DATA_BLOCK "DB_COM_REC_AUX"   // DB37
{ S7_Optimized_Access := 'FALSE' }
VERSION : 0.1
   VAR
      x : Bool;   // Ninguna bomba de intercambiador de soplado en marcha
      x1 : Bool;   // Ninguna bomba de chillers de soplado en marcha
      x2 : Bool;   // Ninguna bomba de intercambiador de envasado en marcha
      x3 : Bool;   // Ninguna bomba de chillers de envasado en marcha
      x4 : Bool;   // Ninguna bomba de torre de enfiamiento de chillers en marcha
      x5 : Bool;   // Ningún Chiller de soplado habilitado
      x6 : Bool;   // Ningún chiller de envasado habilitado
      x7 : Bool;   // Alarma Presente en Chiller de soplado Grande
      x8 : Bool;   // Alarma Presente en Chiller de envasado Grande
      x9 : Bool;   // Chiller de soplado Grande en su máxima capacidad
      x10 : Bool;   // Chiller de envasado Grande en su máxima capacidad
      x11 : Bool;   // Falla Térmico MT007
      x12 : Bool;   // Falla Contactor MT007
      x13 : Bool;   // Falla Térmico MT008
      x14 : Bool;   // Falla Contactor MT008
      x15 : Bool;   // Falla Térmico MT009
      x16 : Bool;   // Falla Contactor MT009
      x17 : Bool;   // Falla Térmico MT010
      x18 : Bool;   // Falla Contactor MT010
      x19 : Bool;   // Falla Térmico MP010
      x20 : Bool;   // Falla Contactor MP010
      x21 : Bool;   // Falla Térmico MP011
      x22 : Bool;   // Falla Contactor MP011
      x23 : Bool;   // Falla Térmico MP012
      x24 : Bool;   // Falla Contactor MP012
      x25 : Bool;   // Falla Térmico MP013
      x26 : Bool;   // Falla Contactor MP013
      x27 : Bool;   // Falla Térmico MP018
      x28 : Bool;   // Falla Contactor MP018
      x29 : Bool;   // Falla Térmico MP019
      x30 : Bool;   // Falla Contactor MP019
      x31 : Bool;   // Falla Térmico V001
      x32 : Bool;   // Falla Contactor V001
      x33 : Bool;   // Falla Térmico V002
      x34 : Bool;   // Falla Contactor V002
      x35 : Bool;   // Falla Térmico V003
      x36 : Bool;   // Falla Contactor V003
      x37 : Bool;   // Falla Térmico MC060
      x38 : Bool;   // Falla Contactor MC060
      x39 : Bool;   // Falla Térmico MC061
      x40 : Bool;   // Falla Contactor MC061
      x41 : Bool;   // Falla Térmico MC062
      x42 : Bool;   // Falla Contactor MC062
      x43 : Bool;   // Falla Térmico MC063
      x44 : Bool;   // Falla Contactor MC063
      x45 : Bool;   // Falla Térmico MC064
      x46 : Bool;   // Falla Contactor MC064
      x47 : Bool;   // Falla Térmico MS050
      x48 : Bool;   // Falla Contactor MS050
      x49 : Bool;   // Falla Térmico MS051
      x50 : Bool;   // Falla Contactor MS051
      x51 : Bool;   // Falla Térmico MS052
      x52 : Bool;   // Falla Contactor MS052
      x53 : Bool;   // Falla Térmico MS053
      x54 : Bool;   // Falla Contactor MS053
      x55 : Bool;   // Falla Presostato Chillers
      x56 : Bool;   // Falla Térmico MS054
      x57 : Bool;   // Falla Contactor MS054
      x58 : Bool;   // Falla Térmico MS055
      x59 : Bool;   // Falla Contactor MS055
      x60 : Bool;   // Falla Térmico MV030
      x61 : Bool;   // Falla Contactor MV030
      x62 : Bool;   // Falla Térmico MV031
      x63 : Bool;   // Falla Contactor MV031
      x64 : Bool;   // Falla Térmico MP014
      x65 : Bool;   // Falla Contactor MP014
      x66 : Bool;   // Falla Térmico MP015
      x67 : Bool;   // Falla Contactor MP015
      x68 : Bool;   // Falla Térmico MC001
      x69 : Bool;   // Falla Contactor MC001
      x70 : Bool;   // Falla Térmico MC002
      x71 : Bool;   // Falla Contactor MC002
      x72 : Bool;   // Falla Térmico MC003
      x73 : Bool;   // Falla Contactor MC003
      x74 : Bool;   // Falla Térmico MC004
      x75 : Bool;   // Falla Contactor MC004
      x76 : Bool;   // Falla Térmico MC005
      x77 : Bool;   // Falla Contactor MC005
      x78 : Bool;   // Falla Flujostato Torres Cavaleto
      x79 : Bool;   // Falla Compresor ABC2 Baja Presion de Aceite
      x80 : Bool;   // Falla Compresor ABC2 Baja Presion de Agua
      x81 : Bool;   // Falla Compresor ABC2 Alta Temperatura de Aire
      x82 : Bool;   // Falla Compresor ABC2 Alta Temperatura de agua
      x83 : Bool;   // Falla Compresor ABC3 Baja Presion de Aceite
      x84 : Bool;   // Falla Compresor ABC3 Baja Presion de Agua
      x85 : Bool;   // Falla Compresor ABC3 Alta Temperatura de Aire
      x86 : Bool;   // Falla Compresor ABC3 Alta Temperatura de agua
      x87 : Bool;   // Falla Compresor ABC4 Baja Presion de Aceite
      x88 : Bool;   // Falla Compresor ABC4 Alta Temperatura de Aire
      x89 : Bool;   // Falla Compresor ABC4 Alta Temperatura de Aire
      x90 : Bool;   // Falla Compresor ABC4 Alta Temperatura de agua
      x91 : Bool;   // Falla Compresor ABC5 Baja Presion de Aceite
      x92 : Bool;   // Falla Compresor ABC5 Alta Temperatura de Aire
      x93 : Bool;   // Falla Compresor ABC5 Alta Temperatura de Aire
      x94 : Bool;   // Falla Compresor ABC5 Alta Temperatura de agua
      x95 : Bool;   // Falla Compresor Bellis & MHW28 Baja Presion Aceite
      x96 : Bool;   // Falla Compresor Bellis & MHW28 Baja Presion de Agua
      x97 : Bool;   // Falla Compresor Bellis & MHW28 Alta temperatura de Aire
      x98 : Bool;   // Falla Compresor Bellis & MHW28 Alta temperatura de Agua
      x99 : Bool;   // Falla Compresor Bellis & MHW28 Falla de Flujostato
      x100 : Bool;   // Requiere Marcha MC001
      x101 : Bool;   // Requiere Marcha MC002
      x102 : Bool;   // Requiere Marcha MC003
      x103 : Bool;   // Requiere Marcha MC004
      x104 : Bool;   // Requiere Marcha MC005
      x105 : Bool;   // Falla Conexión con sensor de Temperatura torres de Cavaleto
      x106 : Bool;   // Falla Conexión con sensor de Temperatura torres de Chillers
      x107 : Bool;   // Falla Conexión con sensor de Presión de ALTA
      x108 : Bool;   // Falla Conexión con sensor de Presión de ALTA redundante
      x109 : Bool;   // Falla Conexión con sensor de Presión de Baja
      x110 : Bool;   // Falla Presión de Alta en Límite Mínimo
      x111 : Bool;   // Falla Presión de Alta en demasiado Baja
      x112 : Bool;   // Falla Presión de Alta en demasiado Alta
      x113 : Bool;   // Falla Presión de Alta en Límite Máximo
      x114 : Bool;   // Falla Presión de Baja en Límite Mínimo
      x115 : Bool;   // Falla Presión de Baja en demasiado Baja
      x116 : Bool;   // Falla Presión de Baja en demasiado Alta
      x117 : Bool;   // Falla Presión de Baja en Límite Máximo
      x118 : Bool;   // Falla en chiller de envasado chico
      x119 : Bool;   // Falla en chiller de soplado chico
      x120 : Bool;   // Horas máximas en Compresor 1
      x121 : Bool;   // Horas máximas en Compresor 2
      x122 : Bool;   // Horas máximas en Compresor 3
      x123 : Bool;   // Horas máximas en Compresor 4
      x124 : Bool;   // Horas máximas en Compresor 5
      x125 : Bool;   // Falla algún contactor en Booster
      x126 : Bool;   // Falla algún guardamotor en Booster
      x127 : Bool;   // Presión Alta en Booster
      x128 : Bool;   // Falla algún contactor en Booster 2
      x129 : Bool;   // Falla algún guardamotor en Booster 2
      x130 : Bool;   // Error lectura analógica Presión Boosters
      x131 : Bool;   // Libre
      x132 : Bool;   // Libre
      x133 : Bool;   // Libre
      x134 : Bool;   // Libre
      x135 : Bool;   // Libre
      x136 : Bool;   // Libre
      x137 : Bool;   // Libre
      x138 : Bool;   // Libre
      x139 : Bool;   // Libre
      x140 : Bool;   // Libre
      x141 : Bool;   // Libre
      x142 : Bool;   // Libre
      x143 : Bool;   // Libre
      x144 : Bool;
      x145 : Bool;
      x146 : Bool;
      x147 : Bool;
      x148 : Bool;
      x149 : Bool;
      x150 : Bool;
      x151 : Bool;
      x152 : Bool;
      x153 : Bool;
      x154 : Bool;
      x155 : Bool;
      x156 : Bool;
      x157 : Bool;
      x158 : Bool;
      x159 : Bool;
      x160 : Bool;
      x161 : Bool;
      x162 : Bool;
      x163 : Bool;
      x164 : Bool;
      x165 : Bool;
      x166 : Bool;
      x167 : Bool;
      x168 : Bool;
      x169 : Bool;
      x170 : Bool;
      x171 : Bool;
      x172 : Bool;
      x173 : Bool;
      x174 : Bool;
      x175 : Bool;
      x176 : Bool;
      x177 : Bool;
      x178 : Bool;
      x179 : Bool;
      x180 : Bool;
      x181 : Bool;
      x182 : Bool;
      x183 : Bool;
      x184 : Bool;
      x185 : Bool;
      x186 : Bool;
      x187 : Bool;
      x188 : Bool;
      x189 : Bool;
      x190 : Bool;
      x191 : Bool;
      x192 : Bool;
      x193 : Bool;
      x194 : Bool;
      x195 : Bool;
      x196 : Bool;
      x197 : Bool;
      x198 : Bool;
      x199 : Bool;
   END_VAR
BEGIN
END_DATA_BLOCK

DATA_BLOCK "DB_BIT_VIDA"   // DB38
{ S7_Optimized_Access := 'FALSE' }
VERSION : 0.1
   VAR
      x : Bool;
      x1 : Bool;
      x2 : Bool;
      x3 : Bool;
      x4 : Bool;
      x5 : Bool;
      x6 : Bool;
      x7 : Bool;
      x8 : Bool;
      x9 : Bool;
      x10 : Bool;
      x11 : Bool;
      x12 : Bool;
      x13 : Bool;
      x14 : Bool;
      x15 : Bool;
      x16 : Bool;
      x17 : Bool;
      x18 : Bool;
      x19 : Bool;
      x20 : Bool;
      x21 : Bool;
      x22 : Bool;
      x23 : Bool;
      x24 : Bool;
      x25 : Bool;
      x26 : Bool;
      x27 : Bool;
      x28 : Bool;
      x29 : Bool;
      x30 : Bool;
      x31 : Bool;
      x32 : Bool;
      x33 : Bool;
      x34 : Bool;
      x35 : Bool;
      x36 : Bool;
      x37 : Bool;
      x38 : Bool;
      x39 : Bool;
      x40 : Bool;
      x41 : Bool;
      x42 : Bool;
      x43 : Bool;
      x44 : Bool;
      x45 : Bool;
      x46 : Bool;
      x47 : Bool;
      x48 : Bool;
      x49 : Bool;
      x50 : Bool;
      x51 : Bool;
      x52 : Bool;
      x53 : Bool;
      x54 : Bool;
      x55 : Bool;
      x56 : Bool;
      x57 : Bool;
      x58 : Bool;
      x59 : Bool;
      x60 : Bool;
      x61 : Bool;
      x62 : Bool;
      x63 : Bool;
      x64 : Bool;
      x65 : Bool;
      x66 : Bool;
      x67 : Bool;
      x68 : Bool;
      x69 : Bool;
      x70 : Bool;
      x71 : Bool;
      x72 : Bool;
      x73 : Bool;
      x74 : Bool;
      x75 : Bool;
      x76 : Bool;
      x77 : Bool;
      x78 : Bool;
      x79 : Bool;
      x80 : Bool;
      x81 : Bool;
      x82 : Bool;
      x83 : Bool;
      x84 : Bool;
      x85 : Bool;
      x86 : Bool;
      x87 : Bool;
      x88 : Bool;
      x89 : Bool;
      x90 : Bool;
      x91 : Bool;
      x92 : Bool;
      x93 : Bool;
      x94 : Bool;
      x95 : Bool;
      x96 : Bool;
      x97 : Bool;
      x98 : Bool;
      x99 : Bool;
      x100 : Bool;
      x101 : Bool;
      x102 : Bool;
      x103 : Bool;
      x104 : Bool;
      x105 : Bool;
      x106 : Bool;
      x107 : Bool;
      x108 : Bool;
      x109 : Bool;
      x110 : Bool;
      x111 : Bool;
      x112 : Bool;
      x113 : Bool;
      x114 : Bool;
      x115 : Bool;
      x116 : Bool;
      x117 : Bool;
      x118 : Bool;
      x119 : Bool;
      x120 : Bool;
      x121 : Bool;
      x122 : Bool;
      x123 : Bool;
      x124 : Bool;
      x125 : Bool;
      x126 : Bool;
      x127 : Bool;
      x128 : Bool;
      x129 : Bool;
      x130 : Bool;
      x131 : Bool;
      x132 : Bool;
      x133 : Bool;
      x134 : Bool;
      x135 : Bool;
      x136 : Bool;
      x137 : Bool;
      x138 : Bool;
      x139 : Bool;
      x140 : Bool;
      x141 : Bool;
      x142 : Bool;
      x143 : Bool;
      x144 : Bool;
      x145 : Bool;
      x146 : Bool;
      x147 : Bool;
      x148 : Bool;
      x149 : Bool;
      x150 : Bool;
      x151 : Bool;
      x152 : Bool;
      x153 : Bool;
      x154 : Bool;
      x155 : Bool;
      x156 : Bool;
      x157 : Bool;
      x158 : Bool;
      x159 : Bool;
      x160 : Bool;
      x161 : Bool;
      x162 : Bool;
      x163 : Bool;
      x164 : Bool;
      x165 : Bool;
      x166 : Bool;
      x167 : Bool;
      x168 : Bool;
      x169 : Bool;
      x170 : Bool;
      x171 : Bool;
      x172 : Bool;
      x173 : Bool;
      x174 : Bool;
      x175 : Bool;
      x176 : Bool;
      x177 : Bool;
      x178 : Bool;
      x179 : Bool;
      x180 : Bool;
      x181 : Bool;
      x182 : Bool;
      x183 : Bool;
      x184 : Bool;
      x185 : Bool;
      x186 : Bool;
      x187 : Bool;
      x188 : Bool;
      x189 : Bool;
      x190 : Bool;
      x191 : Bool;
      x192 : Bool;
      x193 : Bool;
      x194 : Bool;
      x195 : Bool;
      x196 : Bool;
      x197 : Bool;
      x198 : Bool;
      x199 : Bool;
   END_VAR
BEGIN
END_DATA_BLOCK

DATA_BLOCK "AuxiliarAlarmasMTA"   // DB47
{ S7_Optimized_Access := 'FALSE' }
VERSION : 0.1
   VAR
      AlarmaNueva : Bool;   // AlarmaNueva
      AlarmaPresente : Bool;   // AlarmaPresente
      SinAlarmas : Bool;   // SinAlarmas
      Flanco_Bit_Vida : Bool;   // Flanco_Bit_Vida
      Falla_Comunicacion : Bool;   // Falla_Comunicacion
      Bit_Vida_Recibido : Bool;   // Bit_Vida_Recibido
      ReconocerTodas : Bool;   // ReconocerTodas
      Bit_Vida_Enviado : Bool;   // Bit_Vida_Enviado
   END_VAR
BEGIN
END_DATA_BLOCK

DATA_BLOCK "AlarmasDoblePantalla"   // DB86
{ S7_Optimized_Access := 'FALSE' }
VERSION : 0.1
   VAR
      x0 : Bool;   // Ninguna bomba de intercambiador de soplado en marcha
      x1 : Bool;   // Ninguna bomba de chillers de soplado en marcha
      x2 : Bool;   // Ninguna bomba de intercambiador de envasado en marcha
      x3 : Bool;   // Ninguna bomba de chillers de envasado en marcha
      x4 : Bool;   // Ninguna bomba de torre de enfiamiento de chillers en marcha
      x5 : Bool;   // Ningún Chiller de soplado habilitado
      x6 : Bool;   // Ningún chiller de envasado habilitado
      x7 : Bool;   // Alarma Presente en Chiller de soplado Grande
      r0 : Bool;
      r1 : Bool;
      r2 : Bool;
      r3 : Bool;
      r4 : Bool;
      r5 : Bool;
      r6 : Bool;
      r7 : Bool;
      x8 : Bool;   // Alarma Presente en Chiller de envasado Grande
      x9 : Bool;   // Chiller de soplado Grande en su máxima capacidad
      x10 : Bool;   // Chiller de envasado Grande en su máxima capacidad
      x11 : Bool;   // Falla Térmico MT007
      x12 : Bool;   // Falla Contactor MT007
      x13 : Bool;   // Falla Térmico MT008
      x14 : Bool;   // Falla Contactor MT008
      x15 : Bool;   // Falla Térmico MT009
      r8 : Bool;
      r9 : Bool;
      r10 : Bool;
      r11 : Bool;
      r12 : Bool;
      r13 : Bool;
      r14 : Bool;
      r15 : Bool;
      x16 : Bool;   // Falla Contactor MT009
      x17 : Bool;   // Falla Térmico MT010
      x18 : Bool;   // Falla Contactor MT010
      x19 : Bool;   // Falla Térmico MP010
      x20 : Bool;   // Falla Contactor MP010
      x21 : Bool;   // Falla Térmico MP011
      x22 : Bool;   // Falla Contactor MP011
      x23 : Bool;   // Falla Térmico MP012
      r16 : Bool;
      r17 : Bool;
      r18 : Bool;
      r19 : Bool;
      r20 : Bool;
      r21 : Bool;
      r22 : Bool;
      r23 : Bool;
      x24 : Bool;   // Falla Contactor MP012
      x25 : Bool;   // Falla Térmico MP013
      x26 : Bool;   // Falla Contactor MP013
      x27 : Bool;   // Falla Térmico MP018
      x28 : Bool;   // Falla Contactor MP018
      x29 : Bool;   // Falla Térmico MP019
      x30 : Bool;   // Falla Contactor MP019
      x31 : Bool;   // Falla Térmico V001
      r24 : Bool;
      r25 : Bool;
      r26 : Bool;
      r27 : Bool;
      r28 : Bool;
      r29 : Bool;
      r30 : Bool;
      r31 : Bool;
      x32 : Bool;   // Falla Contactor V001
      x33 : Bool;   // Falla Térmico V002
      x34 : Bool;   // Falla Contactor V002
      x35 : Bool;   // Falla Térmico V003
      x36 : Bool;   // Falla Contactor V003
      x37 : Bool;   // Falla Térmico MC060
      x38 : Bool;   // Falla Contactor MC060
      x39 : Bool;   // Falla Térmico MC061
      r32 : Bool;
      r33 : Bool;
      r34 : Bool;
      r35 : Bool;
      r36 : Bool;
      r37 : Bool;
      r38 : Bool;
      r39 : Bool;
      x40 : Bool;   // Falla Contactor MC061
      x41 : Bool;   // Falla Térmico MC062
      x42 : Bool;   // Falla Contactor MC062
      x43 : Bool;   // Falla Térmico MC063
      x44 : Bool;   // Falla Contactor MC063
      x45 : Bool;   // Falla Térmico MC064
      x46 : Bool;   // Falla Contactor MC064
      x47 : Bool;   // Falla Térmico MS050
      r40 : Bool;
      r41 : Bool;
      r42 : Bool;
      r43 : Bool;
      r44 : Bool;
      r45 : Bool;
      r46 : Bool;
      r47 : Bool;
      x48 : Bool;   // Falla Contactor MS050
      x49 : Bool;   // Falla Térmico MS051
      x50 : Bool;   // Falla Contactor MS051
      x51 : Bool;   // Falla Térmico MS052
      x52 : Bool;   // Falla Contactor MS052
      x53 : Bool;   // Falla Térmico MS053
      x54 : Bool;   // Falla Contactor MS053
      x55 : Bool;   // Falla Presostato Chillers
      r48 : Bool;
      r49 : Bool;
      r50 : Bool;
      r51 : Bool;
      r52 : Bool;
      r53 : Bool;
      r54 : Bool;
      r55 : Bool;
      x56 : Bool;   // Falla Térmico MS054
      x57 : Bool;   // Falla Contactor MS054
      x58 : Bool;   // Falla Térmico MS055
      x59 : Bool;   // Falla Contactor MS055
      x60 : Bool;   // Falla Térmico MV030
      x61 : Bool;   // Falla Contactor MV030
      x62 : Bool;   // Falla Térmico MV031
      x63 : Bool;   // Falla Contactor MV031
      r56 : Bool;
      r57 : Bool;
      r58 : Bool;
      r59 : Bool;
      r60 : Bool;
      r61 : Bool;
      r62 : Bool;
      r63 : Bool;
      x64 : Bool;   // Falla Térmico MP014
      x65 : Bool;   // Falla Contactor MP014
      x66 : Bool;   // Falla Térmico MP015
      x67 : Bool;   // Falla Contactor MP015
      x68 : Bool;   // Falla Térmico MC001
      x69 : Bool;   // Falla Contactor MC001
      x70 : Bool;   // Falla Térmico MC002
      x71 : Bool;   // Falla Contactor MC002
      r64 : Bool;
      r65 : Bool;
      r66 : Bool;
      r67 : Bool;
      r68 : Bool;
      r69 : Bool;
      r70 : Bool;
      r71 : Bool;
      x72 : Bool;   // Falla Térmico MC003
      x73 : Bool;   // Falla Contactor MC003
      x74 : Bool;   // Falla Térmico MC004
      x75 : Bool;   // Falla Contactor MC004
      x76 : Bool;   // Falla Térmico MC005
      x77 : Bool;   // Falla Contactor MC005
      x78 : Bool;   // Falla Flujostato Torres Cavaleto
      x79 : Bool;   // Falla Compresor ABC2 Baja Presion de Aceite
      r72 : Bool;
      r73 : Bool;
      r74 : Bool;
      r75 : Bool;
      r76 : Bool;
      r77 : Bool;
      r78 : Bool;
      r79 : Bool;
      x80 : Bool;   // Falla Compresor ABC2 Baja Presion de Agua
      x81 : Bool;   // Falla Compresor ABC2 Alta Temperatura de Aire
      x82 : Bool;   // Falla Compresor ABC2 Alta Temperatura de agua
      x83 : Bool;   // Falla Compresor ABC3 Baja Presion de Aceite
      x84 : Bool;   // Falla Compresor ABC3 Baja Presion de Agua
      x85 : Bool;   // Falla Compresor ABC3 Alta Temperatura de Aire
      x86 : Bool;   // Falla Compresor ABC3 Alta Temperatura de agua
      x87 : Bool;   // Falla Compresor ABC4 Baja Presion de Aceite
      r80 : Bool;
      r81 : Bool;
      r82 : Bool;
      r83 : Bool;
      r84 : Bool;
      r85 : Bool;
      r86 : Bool;
      r87 : Bool;
      x88 : Bool;   // Falla Compresor ABC4 Alta Temperatura de Aire
      x89 : Bool;   // Falla Compresor ABC4 Alta Temperatura de Aire
      x90 : Bool;   // Falla Compresor ABC4 Alta Temperatura de agua
      x91 : Bool;   // Falla Compresor ABC5 Baja Presion de Aceite
      x92 : Bool;   // Falla Compresor ABC5 Alta Temperatura de Aire
      x93 : Bool;   // Falla Compresor ABC5 Alta Temperatura de Aire
      x94 : Bool;   // Falla Compresor ABC5 Alta Temperatura de agua
      x95 : Bool;   // Falla Compresor Bellis & MHW28 Baja Presion Aceite
      r88 : Bool;
      r89 : Bool;
      r90 : Bool;
      r91 : Bool;
      r92 : Bool;
      r93 : Bool;
      r94 : Bool;
      r95 : Bool;
      x96 : Bool;   // Falla Compresor Bellis & MHW28 Baja Presion de Agua
      x97 : Bool;   // Falla Compresor Bellis & MHW28 Alta temperatura de Aire
      x98 : Bool;   // Falla Compresor Bellis & MHW28 Alta temperatura de Agua
      x99 : Bool;   // Falla Compresor Bellis & MHW28 Falla de Flujostato
      x100 : Bool;   // Requiere Marcha MC001
      x101 : Bool;   // Requiere Marcha MC002
      x102 : Bool;   // Requiere Marcha MC003
      x103 : Bool;   // Requiere Marcha MC004
      r96 : Bool;
      r97 : Bool;
      r98 : Bool;
      r99 : Bool;
      r100 : Bool;
      r101 : Bool;
      r102 : Bool;
      r103 : Bool;
      x104 : Bool;   // Requiere Marcha MC005
      x105 : Bool;   // Falla Conexión con sensor de Temperatura torres de Cavaleto
      x106 : Bool;   // Falla Conexión con sensor de Temperatura torres de Chillers
      x107 : Bool;   // Falla Conexión con sensor de Presión de ALTA
      x108 : Bool;   // Falla Conexión con sensor de Presión de ALTA redundante
      x109 : Bool;   // Falla Conexión con sensor de Presión de Baja
      x110 : Bool;   // Falla Presión de Alta en Límite Mínimo
      x111 : Bool;   // Falla Presión de Alta en demasiado Baja
      r104 : Bool;
      r105 : Bool;
      r106 : Bool;
      r107 : Bool;
      r108 : Bool;
      r109 : Bool;
      r110 : Bool;
      r111 : Bool;
      x112 : Bool;   // Falla Presión de Alta en demasiado Alta
      x113 : Bool;   // Falla Presión de Alta en Límite Máximo
      x114 : Bool;   // Falla Presión de Baja en Límite Mínimo
      x115 : Bool;   // Falla Presión de Baja en demasiado Baja
      x116 : Bool;   // Falla Presión de Baja en demasiado Alta
      x117 : Bool;   // Falla Presión de Baja en Límite Máximo
      x118 : Bool;   // Falla en chiller de envasado chico
      x119 : Bool;   // Falla en chiller de soplado chico
      r112 : Bool;
      r113 : Bool;
      r114 : Bool;
      r115 : Bool;
      r116 : Bool;
      r117 : Bool;
      r118 : Bool;
      r119 : Bool;
      x120 : Bool;   // Horas máximas en Compresor 1
      x121 : Bool;   // Horas máximas en Compresor 2
      x122 : Bool;   // Horas máximas en Compresor 3
      x123 : Bool;   // Horas máximas en Compresor 4
      x124 : Bool;   // Horas máximas en Compresor 5
      x125 : Bool;   // Falla algún contactor en Booster 1
      x126 : Bool;   // Falla algún guardamotor en Booster 1
      x127 : Bool;   // Presión Alta en Booster
      r120 : Bool;
      r121 : Bool;
      r122 : Bool;
      r123 : Bool;
      r124 : Bool;
      r125 : Bool;
      r126 : Bool;
      r127 : Bool;
      x128 : Bool;   // Falla algún contactor en Booster 2
      x129 : Bool;   // Falla algún guardamotor en Booster 2
      x130 : Bool;   // Libre
      x131 : Bool;   // Libre
      x132 : Bool;   // Libre
      x133 : Bool;   // Libre
      x134 : Bool;   // Libre
      x135 : Bool;   // Libre
      r128 : Bool;
      r129 : Bool;
      r130 : Bool;
      r131 : Bool;
      r132 : Bool;
      r133 : Bool;
      r134 : Bool;
      r135 : Bool;
      x136 : Bool;   // Libre
      x137 : Bool;   // Libre
      x138 : Bool;   // Libre
      x139 : Bool;   // Libre
      x140 : Bool;   // Libre
      x141 : Bool;   // Libre
      x142 : Bool;   // Libre
      x143 : Bool;   // Libre
      r136 : Bool;
      r137 : Bool;
      r138 : Bool;
      r139 : Bool;
      r140 : Bool;
      r141 : Bool;
      r142 : Bool;
      r143 : Bool;
      x144 : Bool;
      x145 : Bool;
      x146 : Bool;
      x147 : Bool;
      x148 : Bool;
      x149 : Bool;
      x150 : Bool;
      x151 : Bool;
      r144 : Bool;
      r145 : Bool;
      r146 : Bool;
      r147 : Bool;
      r148 : Bool;
      r149 : Bool;
      r150 : Bool;
      r151 : Bool;
      x152 : Bool;
      x153 : Bool;
      x154 : Bool;
      x155 : Bool;
      x156 : Bool;
      x157 : Bool;
      x158 : Bool;
      x159 : Bool;
      r152 : Bool;
      r153 : Bool;
      r154 : Bool;
      r155 : Bool;
      r156 : Bool;
      r157 : Bool;
      r158 : Bool;
      r159 : Bool;
      x160 : Bool;
      x161 : Bool;
      x162 : Bool;
      x163 : Bool;
      x164 : Bool;
      x165 : Bool;
      x166 : Bool;
      x167 : Bool;
      r160 : Bool;
      r161 : Bool;
      r162 : Bool;
      r163 : Bool;
      r164 : Bool;
      r165 : Bool;
      r166 : Bool;
      r167 : Bool;
      x168 : Bool;
      x169 : Bool;
      x170 : Bool;
      x171 : Bool;
      x172 : Bool;
      x173 : Bool;
      x174 : Bool;
      x175 : Bool;
      r168 : Bool;
      r169 : Bool;
      r170 : Bool;
      r171 : Bool;
      r172 : Bool;
      r173 : Bool;
      r174 : Bool;
      r175 : Bool;
      x176 : Bool;
      x177 : Bool;
      x178 : Bool;
      x179 : Bool;
      x180 : Bool;
      x181 : Bool;
      x182 : Bool;
      x183 : Bool;
      r176 : Bool;
      r177 : Bool;
      r178 : Bool;
      r179 : Bool;
      r180 : Bool;
      r181 : Bool;
      r182 : Bool;
      r183 : Bool;
      x184 : Bool;
      x185 : Bool;
      x186 : Bool;
      x187 : Bool;
      x188 : Bool;
      x189 : Bool;
      x190 : Bool;
      x191 : Bool;
      r184 : Bool;
      r185 : Bool;
      r186 : Bool;
      r187 : Bool;
      r188 : Bool;
      r189 : Bool;
      r190 : Bool;
      r191 : Bool;
      x192 : Bool;
      x193 : Bool;
      x194 : Bool;
      x195 : Bool;
      x196 : Bool;
      x197 : Bool;
      x198 : Bool;
      x199 : Bool;
      r192 : Bool;
      r193 : Bool;
      r194 : Bool;
      r195 : Bool;
      r196 : Bool;
      r197 : Bool;
      r198 : Bool;
      r199 : Bool;
   END_VAR
BEGIN
END_DATA_BLOCK

DATA_BLOCK "CFGSirena"   // DB91
{ S7_Optimized_Access := 'FALSE' }
VERSION : 0.1
   VAR
      Motivo1 : Bool;   // Motico 1
      Motivo2 : Bool;   // Motico 2
      Motivo3 : Bool;   // Motico 3
      Motivo4 : Bool;   // Motico 4
      Motivo5 : Bool;   // Motico 5
      Motivo6 : Bool;   // Motico 6
      Motivo7 : Bool;   // Motico 7
      Motivo8 : Bool;   // Motico 8
      Motivo9 : Bool;   // Motico 9
      Motivo10 : Bool;   // Motico 10
      Motivo11 : Bool;   // Motico 11
      Motivo12 : Bool;   // Motico 12
      Motivo13 : Bool;   // Motico 13
      Motivo14 : Bool;   // Motico 14
      Motivo15 : Bool;   // Motico 15
      Motivo16 : Bool;   // Motico 16
      Motivo17 : Bool;   // Motico 17
      Motivo18 : Bool;   // Motico 18
      Motivo19 : Bool;   // Motico 19
      Motivo20 : Bool;   // Motico 20
      Motivo21 : Bool;   // Motico 21
      Motivo22 : Bool;   // Motico 22
      Motivo23 : Bool;   // Motico 23
      Motivo24 : Bool;   // Motico 24
   END_VAR
BEGIN
END_DATA_BLOCK

// folder: Bloques Estándar/Boosters

DATA_BLOCK "Boosters Gral"   // DB62
{ S7_Optimized_Access := 'FALSE' }
VERSION : 0.1
   VAR
      SegBoost1 : Int;   // Segundos acumulados Booster 1
      SegBoost2 : Int;   // Segundos acumulados Booster 2
      MinBoost1 : Int;   // Minutos acumulados booster 1
      MinBoost2 : Int;   // Minutos acumulados booster 2
      HorasBoost1 : DInt;   // Horas acumuladas Boost1
      HorasBoost2 : DInt;   // Horas acumuladas Booster 2
      HorasLim : DInt;   // Horas límite para cambio de prioridad
      TiempoAyudaON_PANEL : Word;   // Tiempo para ayuda Booster Auxiliar PANEL
      TiempoAyudaOFF_PANEL : Word;   // Tiempo para apagar ayuda Booster Auxiliar PANEL
      TiempoAyudaON : S5Time := S5T#1M;   // Tiempo para ayuda Booster Auxiliar
      TiempoAyudaOFF : S5Time := S5T#30S;   // Tiempo para apagar ayuda Booster Auxiliar
      LimArrPrio2 : Real := 8.0e+0;   // Límite para Arranque Booster Prioridad 2
      LimArrPrio1 : Real := 9.0e+0;   // Límite para Arranque Booster Prioridad 1
      LimParPrio2 : Real := 1.1e+1;   // Límite para Parada Booster Prioridad 2
      LimParPrio1 : Real := 1.2e+1;   // Límite para Parada Booster Prioridad 1
      Ctrl_Analogico : Bool;   // Control Boosters por instrumento analógico
   END_VAR
BEGIN
END_DATA_BLOCK

// folder: Compresores/Alta

DATA_BLOCK "AuxiliarVLV"   // DB10
{ S7_Optimized_Access := 'FALSE' }
VERSION : 0.1
   VAR
      DejarAbrirVLV1 : Bool;   // Deja abrir válvula 1
      DejarAbrirVLV2 : Bool;   // Deja abrir válvula 2
      DejarAbrirVLV3 : Bool;   // Deja abrir válvula 3
      DejarAbrirVLV4 : Bool;   // Deja abrir válvula 4
      DejarAbrirVLV5 : Bool;   // Deja abrir válvula 5
      DejarAbrirVLV6 : Bool;
   END_VAR
BEGIN
END_DATA_BLOCK

DATA_BLOCK "DB-PurgaComAlta"   // DB53
{ S7_Optimized_Access := 'FALSE' }
VERSION : 0.1
   VAR
      Habil_PurgaBellis : Bool := true;
      Habil_PurgaABC2 : Bool := true;
      Habil_PurgaABC3 : Bool := true;
      Habil_PurgaABC4 : Bool := true;
      Habil_PurgaABC5 : Bool := true;
      Habil_PurgaABC1 : Bool := true;
      Toff_PurgaBellis : Word := 16#001E;
      Ton_PurgaBellis : Word := 16#001E;
      Toff_PurgaABC2 : Word := 16#001E;
      Ton_PurgaABC2 : Word := 16#001E;
      Toff_PurgaABC3 : Word := 16#001E;
      Ton_PurgaABC3 : Word := 16#001E;
      Toff_PurgaABC4 : Word := 16#001E;
      Ton_PurgaABC4 : Word := 16#001E;
      Toff_PurgaABC5 : Word := 16#001E;
      Ton_PurgaABC5 : Word := 16#001E;
      Toff_PurgaABC1 : Word := 16#001E;
      Ton_PurgaABC1 : Word := 16#001E;
      Prueba_PurgaBellis : Bool;
      Prueba_PurgaABC2 : Bool;
      Prueba_PurgaABC3 : Bool;
      Prueba_PurgaABC4 : Bool;
      Prueba_PurgaABC5 : Bool;
      Prueba_PurgaABC1 : Bool;
   END_VAR
BEGIN
END_DATA_BLOCK

DATA_BLOCK "Agregado Bellis"   // DB63
{ S7_Optimized_Access := 'FALSE' }
VERSION : 0.1
   VAR
      ExcesoTiempo : S5Time := S5T#30M;   // Exceso de tiempo marchando en 1/2 carga
      ForzarCompleta : Bool;   // Forzar carga completa
      QuitarForzado : Bool;   // Quita Forzado de carga completa
      ExcesoTiempoPanel : Int;   // Exceso de tiempo marchando en 1/2 carga desde Panel
   END_VAR
BEGIN
END_DATA_BLOCK

DATA_BLOCK "PanelCompALTA MTA"   // DB75
{ S7_Optimized_Access := 'FALSE' }
VERSION : 0.1
   VAR
      DB_VAR : Int;   // Variable provisional
   END_VAR
BEGIN
END_DATA_BLOCK

DATA_BLOCK "DB-CompAltaDatos"   // DB88
{ S7_Optimized_Access := 'FALSE' }
VERSION : 0.1
   VAR
      Req : Int;   // Cantidad de compresores que hay que encender en total
      F_Osc_1seg : Bool;   // Flanco oscilador período 1 segundo
      MinParGen : Int;   // Minutos de parada general sin requerimiento de ningun compresor
      PanMchCmp1 : Bool;   // Requerimiento de marcha compresor 1
      PanMchCmp2 : Bool;   // Requerimiento de marcha compresor 2
      PanMchCmp3 : Bool;   // Requerimiento de marcha compresor 3
      PanMchCmp4 : Bool;   // Requerimiento de marcha compresor 4
      PanMchCmp5 : Bool;   // Requerimiento de marcha compresor 5
      PanMchCmp6 : Bool;
      TON_ParGen : Bool;   // Timeout estando sin requerimiento de ningun compresor
      TON_ParGen_Lim : Bool;   // Limite excedido Setpoint Timeout estando sin requerimiento de ningun compresor
      ValorParGen : Int := 60;   // Valor actual Timeout estando sin requerimiento de ningun compresor
      Aut1 : Bool;   // Compresor 1 en automático
      Aut2 : Bool;   // Compresor 2 en automático
      Aut3 : Bool;   // Compresor 3 en automático
      Aut4 : Bool;   // Compresor 4 en automático
      Aut5 : Bool;   // Compresor 5 en automático
      Aut6 : Bool;
      TON_ParGenMem : Bool;   // Timeout estando sin requerimiento de ningun compresor memorizado
      CgaPrsCrt : Bool;   // Poner en carga por presion critica
   END_VAR
BEGIN
END_DATA_BLOCK

DATA_BLOCK "FallasCmpALTA"   // DB89
{ S7_Optimized_Access := 'FALSE' }
VERSION : 0.1
   VAR
      FaGen1 : Bool;   // Falla General en tablero 1
      FaGen2 : Bool;   // Falla General en tablero 2
      FaGen3 : Bool;   // Falla General en tablero 3
      FaGen4 : Bool;   // Falla General en tablero 4
      FaGen5 : Bool;   // Falla General en tablero 5
      FaGen6 : Bool;
      FaGen : Bool;   // Falla General
   END_VAR
BEGIN
END_DATA_BLOCK

DATA_BLOCK "CompALTA-MTA"   // DB121
{ S7_Optimized_Access := 'FALSE' }
VERSION : 0.1
   VAR
      FallaGral : Bool;   // Falla General
      FallaCompresor1 : Bool;   // Falla en Compresor 1
      FallaCompresor2 : Bool;   // Falla en Compresor 2
      FallaCompresor3 : Bool;   // Falla en Compresor 3
      FallaCompresor4 : Bool;   // Falla en Compresor 4
      FallaCompresor5 : Bool;   // Falla en Compresor 5
      FallaCompresor6 : Bool;
      EncenderAutoComp1 : Bool;   // Encender automáticamente compresor 1
      EncenderAutoComp2 : Bool;   // Encender automáticamente compresor 2
      EncenderAutoComp3 : Bool;   // Encender automáticamente compresor 3
      EncenderAutoComp4 : Bool;   // Encender automáticamente compresor 4
      EncenderAutoComp5 : Bool;   // Encender automáticamente compresor 5
      EncenderAutoComp6 : Bool;
      IndVCmp1 : Bool;   // Indicación luminosa Verde compresor 1
      IndVCmp2 : Bool;   // Indicación luminosa Verde compresor 2
      IndVCmp3 : Bool;   // Indicación luminosa Verde compresor 3
      IndVCmp4 : Bool;   // Indicación luminosa Verde compresor 4
      IndVCmp5 : Bool;   // Indicación luminosa Verde compresor 5
      IndVCmp6 : Bool;
      IndRCmp1 : Bool;   // Indicación luminosa Roja Compresor 1
      IndRCmp2 : Bool;   // Indicación luminosa Roja Compresor 2
      IndRCmp3 : Bool;   // Indicación luminosa Roja Compresor 3
      IndRCmp4 : Bool;   // Indicación luminosa Roja Compresor 4
      IndRCmp5 : Bool;   // Indicación luminosa Roja Compresor 5
      IndRCmp6 : Bool;
      CmpReq : Word;   // Cantidad de compresores de alta requeridos
      IndMarchaCmp1 : Bool;   // Indicador marcha Compresor1
      IndMarchaCmp2 : Bool;   // Indicador marcha Compresor2
      IndMarchaCmp3 : Bool;   // Indicador marcha Compresor3
      IndMarchaCmp4 : Bool;   // Indicador marcha Compresor4
      IndMarchaCmp5 : Bool;   // Indicador marcha Compresor5
      IndMarchaCmp6 : Bool;
      OvrLimP1 : Bool;   // Compresor 1 sobre el límite de presión superior
      OvrLimP2 : Bool;   // Compresor 2 sobre el límite de presión superior
      OvrLimP3 : Bool;   // Compresor 3 sobre el límite de presión superior
      OvrLimP4 : Bool;   // Compresor 4 sobre el límite de presión superior
      OvrLimP5 : Bool;   // Compresor 5 sobre el límite de presión superior
      OvrLimP6 : Bool;
      UndLimP1 : Bool;   // Compresor 1 por debajo del límite de presión inferior
      RESETPrioridades : Bool;   // Reset de Prioridades
      UndLimP2 : Bool;   // Compresor 2 por debajo del límite de presión inferior
      UndLimP3 : Bool;   // Compresor 3 por debajo del límite de presión inferior
      UndLimP4 : Bool;   // Compresor 4 por debajo del límite de presión inferior
      UndLimP5 : Bool;   // Compresor 5 por debajo del límite de presión inferior
      UndLimP6 : Bool;
      PrsMed : Real;   // Presión media expresada como número real
      MchP1 : Bool;   // Marchar compresor de Prioridad 1
      MchP2 : Bool;   // Marchar compresor de Prioridad 2
      MchP3 : Bool;   // Marchar compresor de Prioridad 3
      MchP4 : Bool;   // Marchar compresor de Prioridad 4
      MchP5 : Bool;   // Marchar compresor de Prioridad 5
      MchP6 : Bool;
      CgaP1 : Bool;   // Poner en carga Prioridad 1
      CgaP2 : Bool;   // Poner en carga Prioridad 2
      CgaP3 : Bool;   // Poner en carga Prioridad 3
      CgaP4 : Bool;   // Poner en carga Prioridad 4
      CgaP5 : Bool;   // Poner en carga Prioridad 5
      CgaP6 : Bool;
      VRealCmp1 : Int;   // Nro de Prioridad real del compresor 1
      Reserva : Int;
      VRealCmp2 : Int;   // Nro de Prioridad real del compresor 2
      Reserva1 : Int;
      VRealCmp3 : Int;   // Nro de Prioridad real del compresor 3
      Reserva2 : Int;
      VRealCmp4 : Int;   // Nro de Prioridad real del compresor 4
      Reserva3 : Int;
      VRealCmp5 : Int;   // Nro de Prioridad real del compresor 5
      Reserva4 : Int;
      VRealCmp6 : Int;
      Reserva5 : Int;
      ReqMch1 : Bool;   // Requerir Marcha de compresor 1
      ReqMch2 : Bool;   // Requerir Marcha de compresor 2
      ReqMch3 : Bool;   // Requerir Marcha de compresor 3
      ReqMch4 : Bool;   // Requerir Marcha de compresor 4
      ReqMch5 : Bool;   // Requerir Marcha de compresor 5
      ReqMch6 : Bool;
      SinReq1 : Bool;   // Compresor 1 Sin requerimiento
      SinReq2 : Bool;   // Compresor 2 Sin requerimiento
      SinReq3 : Bool;   // Compresor 3 Sin requerimiento
      SinReq4 : Bool;   // Compresor 4 Sin requerimiento
      SinReq5 : Bool;   // Compresor 5 Sin requerimiento
      SinReq6 : Bool;
      ManP1 : Bool;   // Prioridad 1 en Manual
      ManP2 : Bool;   // Prioridad 2 en Manual
      ManP3 : Bool;   // Prioridad 3 en Manual
      ManP4 : Bool;   // Prioridad 4 en Manual
      ManP5 : Bool;   // Prioridad 5 en Manual
      ManP6 : Bool;
      CicloIni : Bool;   // Ciclo inicial
      ReqCga1 : Bool;   // Se Necesita poner en carga
      ReqCga2 : Bool;   // Se Necesita poner en carga
      ReqCga3 : Bool;   // Se Necesita poner en carga
      ReqCga4 : Bool;   // Se Necesita poner en carga
      ReqCga5 : Bool;   // Se Necesita poner en carga
      ReqCga6 : Bool;
      ReqCrr : Int;   // Requerimiento inicial corregido
      AnimCMP1 : Int;   // Word Animación Compresor 1
      AnimCMP2 : Int;   // Word Animación Compresor 2
      AnimCMP3 : Int;   // Word Animación Compresor 3
      AnimCMP4 : Int;   // Word Animación Compresor 4
      AnimCMP5 : Int;   // Word Animación Compresor 5
      AnimCMP6 : Int;
      AnimGen : Int;   // Word Animación Maq Est General
      Reset : Bool;   // Reset
      UltPriDis : Int;   // Guarda valor de última prioridad que tenía un compresor disponible
      CntReqIte : Int;   // Cantidad de compresores según las iteraciones realizadas
      CntReqCrr : Int;   // Requerimiento inicial corregido
      CntCmpDisp : Int;   // acumula cantidad compresores disponibles hasta alcanzar numero requerido
      IndVP1 : Bool;   // Indicador Verde con parpadeo 1
      IndVP2 : Bool;   // Indicador Verde con parpadeo 2
      IndVP3 : Bool;   // Indicador Verde con parpadeo 3
      IndVP4 : Bool;   // Indicador Verde con parpadeo 4
      IndVP5 : Bool;   // Indicador Verde con parpadeo 5
      IndVP6 : Bool;
      OvrLimPCRT : Bool;   // Sobre límite de presión crítica superior
      UndLimPCRT : Bool;   // Debajo del límite de presión crítica inferior
   END_VAR
BEGIN
END_DATA_BLOCK

DATA_BLOCK "DBParamCmpALTA-MTA"   // DB122
{ S7_Optimized_Access := 'FALSE' }
VERSION : 0.1
   VAR
      LimSupP1 : Real := 42.0;   // Límite Superior para regulación 1
      LimSupP2 : Real := 41.5;   // Límite Superior para regulación 2
      LimSupP3 : Real := 41.0;   // Límite Superior para regulación 3
      LimSupP4 : Real := 40.5;   // Límite Superior para regulación 4
      LimSupP5 : Real := 40.0;   // Límite Superior para regulación 5
      LimSupP6 : Real := 39.5;
      LimInfP1 : Real := 41.5;   // Límite Inferior para regulación 1
      LimInfP2 : Real := 41.0;   // Límite Inferior para regulación 2
      LimInfP3 : Real := 40.5;   // Límite Inferior para regulación 3
      LimInfP4 : Real := 40.0;   // Límite Inferior para regulación 4
      LimInfP5 : Real := 39.5;   // Límite Inferior para regulación 5
      LimInfP6 : Real := 39.0;
      DelPrs : Real := 0.0;   // Separación entre presiones de un compresor a otro
      HstPrs : Real := 0.5;   // Histeresis para límites de presión
      PrsMax : Real := 42.0;   // Presión superior del compresor con máxima prioridad
      HstPrsCrt : Real := 1.0;   // Histeresis para presión crítica
      LimSupPCRT : Real := 39.0;   // Límite Superior Presión Crítica
      LimInfPCRT : Real := 38.0;   // Límite Inferior Presión Crítica
      LMedia1 : Real := 41.75;   // Limite Superior para Bellis en prioridad 1
      LMedia2 : Real := 41.25;   // Limite Superior para Bellis en prioridad 2
      LMedia3 : Real := 40.75;   // Limite Superior para Bellis en prioridad 3
      LMedia4 : Real := 40.25;   // Limite Superior para Bellis en prioridad 4
      LMedia5 : Real := 39.75;   // Limite Superior para Bellis en prioridad 5
      LMedia6 : Real := 39.25;
      MediaHist : Real := 0.25;   // Mitad de la excursión de presión
      TempCritEnclav : Real := 50.0;
   END_VAR
BEGIN
END_DATA_BLOCK

DATA_BLOCK "DBTiemposCmpAltaMTA"   // DB123
{ S7_Optimized_Access := 'FALSE' }
VERSION : 0.1
   VAR
      FNueReqIni : Bool;   // El valor de requerimiento de compresores iniciales ha cambiado
      Reserva2 : Bool;
      Reserva3 : Bool;
      Reserva4 : Bool;
      Reserva5 : Bool;
      TVAC : S5Time := S5T#1H;   // Tiempo en vacío
      TVACPANEL : Int := 60;   // Tiempo en vacío desde Panel
      TVACPEsc : Int := 60;   // Tiempo en vacío desde Panel Escalado
      RetSinRec : S5Time := S5T#1H;   // Tiempo sin requerimiento
      RetSinRecPANEL : Int := 60;   // Tiempo sin requerimiento desde Panel
      RetSinRecPEsc : Int := 60;   // Tiempo sin requerimiento desde Panel Escalado
   END_VAR
BEGIN
END_DATA_BLOCK

DATA_BLOCK "Sopladoras"   // DB124
{ S7_Optimized_Access := 'FALSE' }
VERSION : 0.1
   VAR
      Sop1 : Bool;   // Sopladora 1 en marcha
      Sop2 : Bool;   // Sopladora 2 en marcha
      Sop3 : Bool;   // Sopladora 3 en marcha
      TStopSop : S5Time := S5T#1H;   // Tiempo de parada para Sopladora
      TStopSopPanel : Int := 60;   // Tiempo de parada para Sopladora desde Panel
      NinSOP : Bool;   // Ninguna Sopladora
      ReqSp1 : Int;   // Cantidad de compresores Requeridos para Sopladora 1
      ReqSp2 : Int;   // Cantidad de compresores Requeridos para Sopladora 2
      ReqSp3 : Int;   // Cantidad de compresores Requeridos para Sopladora 3
      ReqIni : Int;   // Cantidad de compresores requeridos solo por sopladoras
      FinClcReq : Bool;   // Finalizar calculo de compresores requeridos
   END_VAR
BEGIN
END_DATA_BLOCK

DATA_BLOCK "DB-PrioridadesCmpAlta"   // DB125
{ S7_Optimized_Access := 'FALSE' }
VERSION : 0.1
   VAR
      Vcmp0 : Int;   // Nro de prioridad del compresor 0 desde panel
      Vcmp1 : Int := 1;   // Nro de prioridad del compresor 1 desde panel
      Vcmp2 : Int := 2;   // Nro de prioridad del compresor 2 desde panel
      Vcmp3 : Int := 3;   // Nro de prioridad del compresor 3 desde panel
      Vcmp4 : Int := 4;   // Nro de prioridad del compresor 4 desde panel
      Vcmp5 : Int := 5;   // Nro de prioridad del compresor 5 desde panel
      Vcmp6 : Int;
      fDecPri1 : Bool;   // Flanco decrementar prioridad compresor 1
      fDecPri2 : Bool;   // Flanco decrementar prioridad compresor 2
      fDecPri3 : Bool;   // Flanco decrementar prioridad compresor 3
      fDecPri4 : Bool;   // Flanco decrementar prioridad compresor 4
      fDecPri5 : Bool;   // Flanco decrementar prioridad compresor 5
      fDecPri6 : Bool;
      fIncPri1 : Bool;   // Flanco incrementar prioridad compresor 1
      fIncPri2 : Bool;   // Flanco incrementar prioridad compresor 2
      fIncPri3 : Bool;   // Flanco incrementar prioridad compresor 3
      fIncPri4 : Bool;   // Flanco incrementar prioridad compresor 4
      fIncPri5 : Bool;   // Flanco incrementar prioridad compresor 5
      fIncPri6 : Bool;
      IncPri1 : Bool;   // Incrementar prioridad compresor 1
      IncPri2 : Bool;   // Incrementar prioridad compresor 2
      IncPri3 : Bool;   // Incrementar prioridad compresor 3
      IncPri4 : Bool;   // Incrementar prioridad compresor 4
      IncPri5 : Bool;   // Incrementar prioridad compresor 5
      IncPri6 : Bool;
      DecPri1 : Bool;   // Decrementar prioridad compresor 1
      DecPri2 : Bool;   // Decrementar prioridad compresor 2
      DecPri3 : Bool;   // Decrementar prioridad compresor 3
      DecPri4 : Bool;   // Decrementar prioridad compresor 4
      DecPri5 : Bool;   // Decrementar prioridad compresor 5
      DecPri6 : Bool;
   END_VAR
BEGIN
END_DATA_BLOCK

DATA_BLOCK "DB-AccionamientosCmpAlta"   // DB126
{ S7_Optimized_Access := 'FALSE' }
VERSION : 0.1
   VAR
      DB_VAR : Int;   // Variable provisional
   END_VAR
BEGIN
END_DATA_BLOCK

DATA_BLOCK "PanelCmpAlta"   // DB135
{ S7_Optimized_Access := 'FALSE' }
VERSION : 0.1
   VAR
      AnimMenu1 : Int;   // Animación Menu Mc001
      AnimMenu2 : Int;   // Animación Menu Mc002
      AnimMenu3 : Int;   // Animación Menu Mc003
      AnimMenu4 : Int;   // Animación Menu Mc004
      AnimMenu5 : Int;   // Animación Menu Mc005
      AnimMenu6 : Int;
      SPON1 : Real;   // SetPoint Manual MC001
      SPON2 : Real;   // SetPoint Manual MC002
      SPON3 : Real;   // SetPoint Manual MC003
      SPON4 : Real;   // SetPoint Manual MC004
      SPON5 : Real;   // SetPoint Manual MC005
      SPON6 : Real;
      SPOFF1 : Real;   // SetPoint Manual MC001
      SPOFF2 : Real;   // SetPoint Manual MC002
      SPOFF3 : Real;   // SetPoint Manual MC003
      SPOFF4 : Real;   // SetPoint Manual MC004
      SPOFF5 : Real;   // SetPoint Manual MC005
      SPOFF6 : Real;
      MantMC001 : Bool;   // Mantenimiento MC001
      MantMC002 : Bool;   // Mantenimiento MC002
      MantMC003 : Bool;   // Mantenimiento MC003
      MantMC004 : Bool;   // Mantenimiento MC004
      MantMC005 : Bool;   // Mantenimiento MC005
      MantMC006 : Bool;
      MachaMC001 : Bool;   // Orden de Marcha para MC001
      MachaMC002 : Bool;   // Orden de Marcha para MC002
      MachaMC003 : Bool;   // Orden de Marcha para MC003
      MachaMC004 : Bool;   // Orden de Marcha para MC004
      MachaMC005 : Bool;   // Orden de Marcha para MC005
      MachaMC006 : Bool;
      MarchaPanelMC001 : Bool;   // Pulsador Marcha Panel MC001
      MarchaPanelMC002 : Bool;   // Pulsador Marcha Panel MC002
      MarchaPanelMC003 : Bool;   // Pulsador Marcha Panel MC003
      MarchaPanelMC004 : Bool;   // Pulsador Marcha Panel MC004
      MarchaPanelMC005 : Bool;   // Pulsador Marcha Panel MC005
      MarchaPanelMC006 : Bool;
      ParadaPanelMC001 : Bool;   // Pulsador Parada Panel MC001
      ParadaPanelMC002 : Bool;   // Pulsador Parada Panel MC002
      ParadaPanelMC003 : Bool;   // Pulsador Parada Panel MC003
      ParadaPanelMC004 : Bool;   // Pulsador Parada Panel MC004
      ParadaPanelMC005 : Bool;   // Pulsador Parada Panel MC005
      ParadaPanelMC006 : Bool;
      MediaCargaBellis : Bool;   // Compresor Bellis Media Carga
      AbrirVLV1 : Bool;   // Abrir Válvula 1
      AbrirVLV2 : Bool;   // Abrir Válvula 2
      AbrirVLV3 : Bool;   // Abrir Válvula 3
      AbrirVLV4 : Bool;   // Abrir Válvula 4
      AbrirVLV5 : Bool;   // Abrir Válvula 5
      AbrirVLV6 : Bool;
      AbrirVLV3b : Bool;   // Abrir Válvula 3b
   END_VAR
BEGIN
END_DATA_BLOCK

DATA_BLOCK "ModoManualCompAlta"   // DB136
{ S7_Optimized_Access := 'FALSE' }
VERSION : 0.1
   VAR
      MarchaFPanel1 : Bool;   // Orden de forzar Marcha desde el panel MC001
      MarchaFPanel2 : Bool;   // Orden de forzar Marcha desde el panel MC002
      MarchaFPanel3 : Bool;   // Orden de forzar Marcha desde el panel MC003
      MarchaFPanel4 : Bool;   // Orden de forzar Marcha desde el panel MC004
      MarchaFPanel5 : Bool;   // Orden de forzar Marcha desde el panel MC005
      MarchaFPanel6 : Bool;
      ParadaFPanel1 : Bool;   // Orden de forzar Parada desde el panel MC001
      ParadaFPanel2 : Bool;   // Orden de forzar Parada desde el panel MC002
      ParadaFPanel3 : Bool;   // Orden de forzar Parada desde el panel MC003
      ParadaFPanel4 : Bool;   // Orden de forzar Parada desde el panel MC004
      ParadaFPanel5 : Bool;   // Orden de forzar Parada desde el panel MC005
      ParadaFPanel6 : Bool;
      OrdenMarchaForzada1 : Bool;   // Orden de Marcha Forzada MC001
      OrdenMarchaForzada2 : Bool;   // Orden de Marcha Forzada MC002
      OrdenMarchaForzada3 : Bool;   // Orden de Marcha Forzada MC003
      OrdenMarchaForzada4 : Bool;   // Orden de Marcha Forzada MC004
      OrdenMarchaForzada5 : Bool;   // Orden de Marcha Forzada MC005
      OrdenMarchaForzada6 : Bool;
      VlvManual1 : Bool;   // Válvula manual MC001
      VlvManual2 : Bool;   // Válvula manual MC002
      VlvManual3 : Bool;   // Válvula manual MC003
      VlvManual4 : Bool;   // Válvula manual MC004
      VlvManual5 : Bool;   // Válvula manual MC005
      VlvManual6 : Bool;
      SPON1 : Real;   // Setpoint arranque MC001
      SPON2 : Real;   // Setpoint arranque MC002
      SPON3 : Real;   // Setpoint arranque MC003
      SPON4 : Real;   // Setpoint arranque MC004
      SPON5 : Real;   // Setpoint arranque MC005
      SPON6 : Real;
      SPOFF1 : Real;   // Setpoint parada MC001
      SPOFF2 : Real;   // Setpoint parada MC002
      SPOFF3 : Real;   // Setpoint parada MC003
      SPOFF4 : Real;   // Setpoint parada MC004
      SPOFF5 : Real;   // Setpoint parada MC005
      SPOFF6 : Real;
      SPON3b : Real;   // Setpoint arranque b MC003
      SPOFF3b : Real;   // Setpoint parada b MC003
      VlvManual3b : Bool;   // Válvula manual MC003b
   END_VAR
BEGIN
END_DATA_BLOCK

// folder: Compresores/Alta/Máquina de Estados

DATA_BLOCK "EstadosCmpALTA-MTA"   // DB120
{ S7_Optimized_Access := 'FALSE' }